// TIA Portal project "uppgift2" (V18) (continued)
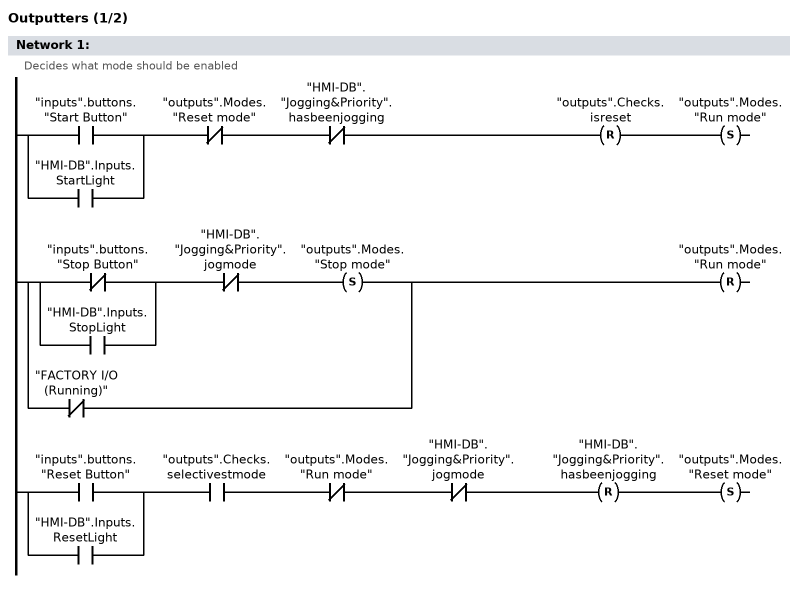
   RUNG wire#powerrail
      Contact( "inputs".buttons."Start Button" )
      wire#w1
      I_Contact( "outputs".Modes."Reset mode" )
      I_Contact( "HMI-DB"."Jogging&Priority".hasbeenjogging )
      R_Coil( "outputs".Checks.isreset )
      S_Coil( "outputs".Modes."Run mode" )
   END_RUNG
   RUNG wire#powerrail
      Contact( "HMI-DB".Inputs.StartLight )
   END_RUNG wire#w1
   RUNG wire#powerrail
      I_Contact( "inputs".buttons."Stop Button" )
      wire#w2
      I_Contact( "HMI-DB"."Jogging&Priority".jogmode )
      S_Coil( "outputs".Modes."Stop mode" )
      wire#w3
      R_Coil( "outputs".Modes."Run mode" )
   END_RUNG
   RUNG wire#powerrail
      Contact( "HMI-DB".Inputs.StopLight )
   END_RUNG wire#w2
   RUNG wire#powerrail
      I_Contact( "FACTORY I/O (Running)" )
   END_RUNG wire#w3
   RUNG wire#powerrail
      Contact( "inputs".buttons."Reset Button" )
      wire#w4
      Contact( "outputs".Checks.selectivestmode )
      I_Contact( "outputs".Modes."Run mode" )
      I_Contact( "HMI-DB"."Jogging&Priority".jogmode )
      R_Coil( "HMI-DB"."Jogging&Priority".hasbeenjogging )
      S_Coil( "outputs".Modes."Reset mode" )
   END_RUNG
   RUNG wire#powerrail
      Contact( "HMI-DB".Inputs.ResetLight )
   END_RUNG wire#w4
   // the same network as SCL:
   IF ("inputs".buttons."Start Button" OR "HMI-DB".Inputs.StartLight) AND NOT "outputs".Modes."Reset mode" AND NOT "HMI-DB"."Jogging&Priority".hasbeenjogging THEN
       "outputs".Checks.isreset := FALSE;
       "outputs".Modes."Run mode" := TRUE;
   END_IF;
   #_w1 := (NOT "inputs".buttons."Stop Button" OR "HMI-DB".Inputs.StopLight) AND NOT "HMI-DB"."Jogging&Priority".jogmode;
   IF #_w1 THEN "outputs".Modes."Stop mode" := TRUE; END_IF;
   IF #_w1 OR NOT "FACTORY I/O (Running)" THEN "outputs".Modes."Run mode" := FALSE; END_IF;
   IF ("inputs".buttons."Reset Button" OR "HMI-DB".Inputs.ResetLight) AND "outputs".Checks.selectivestmode AND NOT "outputs".Modes."Run mode" AND NOT "HMI-DB"."Jogging&Priority".jogmode THEN
       "HMI-DB"."Jogging&Priority".hasbeenjogging := FALSE;
       "outputs".Modes."Reset mode" := TRUE;
   END_IF;
END_REGION

REGION Network 2
   // Turns on the acutators if the correct signal is on
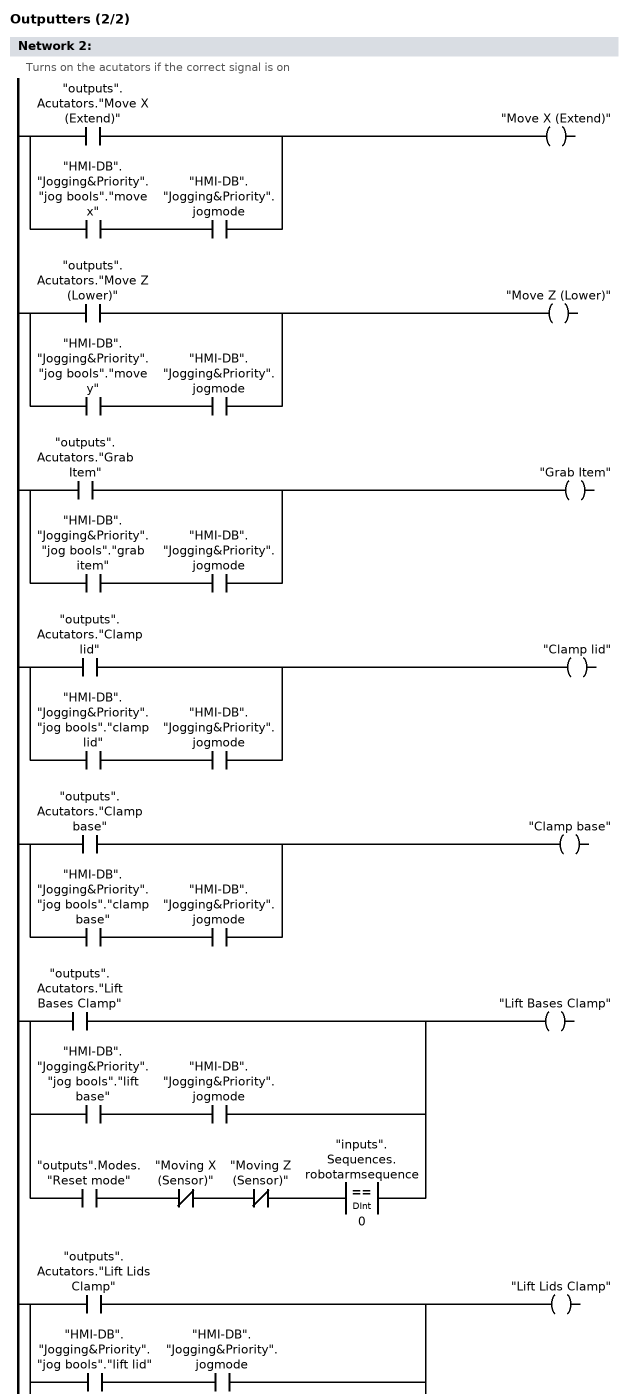
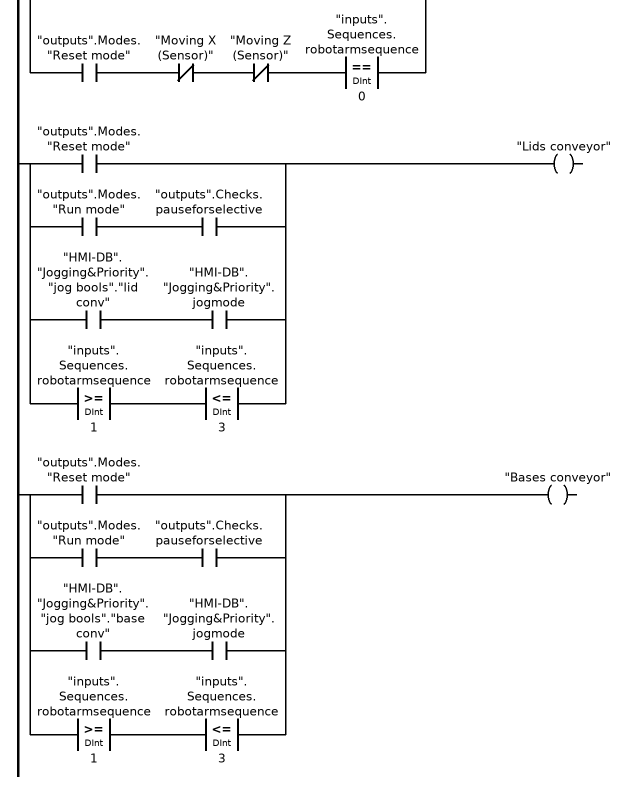
   RUNG wire#powerrail
      Contact( "outputs".Acutators."Move X (Extend)" )
      wire#w1
      Coil( "Move X (Extend)" )
   END_RUNG
   RUNG wire#powerrail
      Contact( "HMI-DB"."Jogging&Priority"."jog bools"."move x" )
      Contact( "HMI-DB"."Jogging&Priority".jogmode )
   END_RUNG wire#w1
   RUNG wire#powerrail
      Contact( "outputs".Acutators."Move Z (Lower)" )
      wire#w2
      Coil( "Move Z (Lower)" )
   END_RUNG
   RUNG wire#powerrail
      Contact( "HMI-DB"."Jogging&Priority"."jog bools"."move y" )
      Contact( "HMI-DB"."Jogging&Priority".jogmode )
   END_RUNG wire#w2
   RUNG wire#powerrail
      Contact( "outputs".Acutators."Grab Item" )
      wire#w3
      Coil( "Grab Item" )
   END_RUNG
   RUNG wire#powerrail
      Contact( "HMI-DB"."Jogging&Priority"."jog bools"."grab item" )
      Contact( "HMI-DB"."Jogging&Priority".jogmode )
   END_RUNG wire#w3
   RUNG wire#powerrail
      Contact( "outputs".Acutators."Clamp lid" )
      wire#w4
      Coil( "Clamp lid" )
   END_RUNG
   RUNG wire#powerrail
      Contact( "HMI-DB"."Jogging&Priority"."jog bools"."clamp lid" )
      Contact( "HMI-DB"."Jogging&Priority".jogmode )
   END_RUNG wire#w4
   RUNG wire#powerrail
      Contact( "outputs".Acutators."Clamp base" )
      wire#w5
      Coil( "Clamp base" )
   END_RUNG
   RUNG wire#powerrail
      Contact( "HMI-DB"."Jogging&Priority"."jog bools"."clamp base" )
      Contact( "HMI-DB"."Jogging&Priority".jogmode )
   END_RUNG wire#w5
   RUNG wire#powerrail
      Contact( "outputs".Acutators."Lift Bases Clamp" )
      wire#w6
      Coil( "Lift Bases Clamp" )
   END_RUNG
   RUNG wire#powerrail
      Contact( "HMI-DB"."Jogging&Priority"."jog bools"."lift base" )
      Contact( "HMI-DB"."Jogging&Priority".jogmode )
   END_RUNG wire#w6
   RUNG wire#powerrail
      Contact( "outputs".Modes."Reset mode" )
      I_Contact( "Moving X (Sensor)" )
      I_Contact( "Moving Z (Sensor)" )
      { S7_Templates := "SrcType := DInt" } EQ_Contact(in1 := "inputs".Sequences.robotarmsequence, in2 := 0)
   END_RUNG wire#w6
   RUNG wire#powerrail
      Contact( "outputs".Acutators."Lift Lids Clamp" )
      wire#w7
      Coil( "Lift Lids Clamp" )
   END_RUNG
   RUNG wire#powerrail
      Contact( "HMI-DB"."Jogging&Priority"."jog bools"."lift lid" )
      Contact( "HMI-DB"."Jogging&Priority".jogmode )
   END_RUNG wire#w7
   RUNG wire#powerrail
      Contact( "outputs".Modes."Reset mode" )
      I_Contact( "Moving X (Sensor)" )
      I_Contact( "Moving Z (Sensor)" )
      { S7_Templates := "SrcType := DInt" } EQ_Contact(in1 := "inputs".Sequences.robotarmsequence, in2 := 0)
   END_RUNG wire#w7
   RUNG wire#powerrail
      Contact( "outputs".Modes."Reset mode" )
      wire#w8
      Coil( "Lids conveyor" )
   END_RUNG
   RUNG wire#powerrail
      Contact( "outputs".Modes."Run mode" )
      Contact( "outputs".Checks.pauseforselective )
   END_RUNG wire#w8
   RUNG wire#powerrail
      Contact( "HMI-DB"."Jogging&Priority"."jog bools"."lid conv" )
      Contact( "HMI-DB"."Jogging&Priority".jogmode )
   END_RUNG wire#w8
   RUNG wire#powerrail
      { S7_Templates := "SrcType := DInt" } GE_Contact(in1 := "inputs".Sequences.robotarmsequence, in2 := 1)
      { S7_Templates := "SrcType := DInt" } LE_Contact(in1 := "inputs".Sequences.robotarmsequence, in2 := 3)
   END_RUNG wire#w8
   RUNG wire#powerrail
      Contact( "outputs".Modes."Reset mode" )
      wire#w9
      Coil( "Bases conveyor" )
   END_RUNG
   RUNG wire#powerrail
      Contact( "outputs".Modes."Run mode" )
      Contact( "outputs".Checks.pauseforselective )
   END_RUNG wire#w9
   RUNG wire#powerrail
      Contact( "HMI-DB"."Jogging&Priority"."jog bools"."base conv" )
      Contact( "HMI-DB"."Jogging&Priority".jogmode )
   END_RUNG wire#w9
   RUNG wire#powerrail
      { S7_Templates := "SrcType := DInt" } GE_Contact(in1 := "inputs".Sequences.robotarmsequence, in2 := 1)
      { S7_Templates := "SrcType := DInt" } LE_Contact(in1 := "inputs".Sequences.robotarmsequence, in2 := 3)
   END_RUNG wire#w9
   // the same network as SCL:
   "Move X (Extend)" := "outputs".Acutators."Move X (Extend)" OR ("HMI-DB"."Jogging&Priority"."jog bools"."move x" AND "HMI-DB"."Jogging&Priority".jogmode);
   "Move Z (Lower)" := "outputs".Acutators."Move Z (Lower)" OR ("HMI-DB"."Jogging&Priority"."jog bools"."move y" AND "HMI-DB"."Jogging&Priority".jogmode);
   "Grab Item" := "outputs".Acutators."Grab Item" OR ("HMI-DB"."Jogging&Priority"."jog bools"."grab item" AND "HMI-DB"."Jogging&Priority".jogmode);
   "Clamp lid" := "outputs".Acutators."Clamp lid" OR ("HMI-DB"."Jogging&Priority"."jog bools"."clamp lid" AND "HMI-DB"."Jogging&Priority".jogmode);
   "Clamp base" := "outputs".Acutators."Clamp base" OR ("HMI-DB"."Jogging&Priority"."jog bools"."clamp base" AND "HMI-DB"."Jogging&Priority".jogmode);
   "Lift Bases Clamp" := "outputs".Acutators."Lift Bases Clamp" OR ("HMI-DB"."Jogging&Priority"."jog bools"."lift base" AND "HMI-DB"."Jogging&Priority".jogmode) OR ("outputs".Modes."Reset mode" AND NOT "Moving X (Sensor)" AND NOT "Moving Z (Sensor)" AND ("inputs".Sequences.robotarmsequence = 0));
   "Lift Lids Clamp" := "outputs".Acutators."Lift Lids Clamp" OR ("HMI-DB"."Jogging&Priority"."jog bools"."lift lid" AND "HMI-DB"."Jogging&Priority".jogmode) OR ("outputs".Modes."Reset mode" AND NOT "Moving X (Sensor)" AND NOT "Moving Z (Sensor)" AND ("inputs".Sequences.robotarmsequence = 0));
   "Lids conveyor" := "outputs".Modes."Reset mode" OR ("outputs".Modes."Run mode" AND "outputs".Checks.pauseforselective) OR ("HMI-DB"."Jogging&Priority"."jog bools"."lid conv" AND "HMI-DB"."Jogging&Priority".jogmode) OR (("inputs".Sequences.robotarmsequence >= 1) AND ("inputs".Sequences.robotarmsequence <= 3));
   "Bases conveyor" := "outputs".Modes."Reset mode" OR ("outputs".Modes."Run mode" AND "outputs".Checks.pauseforselective) OR ("HMI-DB"."Jogging&Priority"."jog bools"."base conv" AND "HMI-DB"."Jogging&Priority".jogmode) OR (("inputs".Sequences.robotarmsequence >= 1) AND ("inputs".Sequences.robotarmsequence <= 3));
END_REGION
END_FUNCTION

// folder: lids/bases

FUNCTION "lids" : Void   // FC3, LAD
{ S7_Optimized_Access := 'TRUE' }
VERSION : 0.1
// Controls the lid clamp and lift and controls when the robots sequence should start
   VAR_TEMP   // added for the SCL form of the ladder/FBD networks
      _w1 : Bool;
   END_VAR
BEGIN

REGION Network 1
   // Runs the emitter if sequence is 0 and lids vision doesnt detect any lid
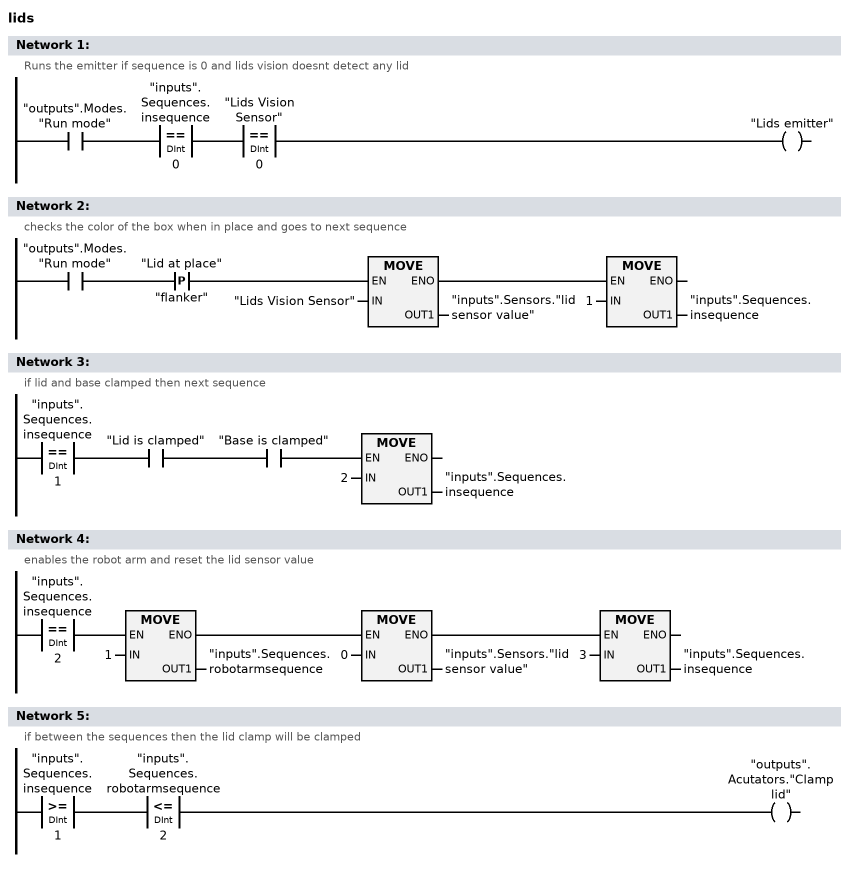
   RUNG wire#powerrail
      Contact( "outputs".Modes."Run mode" )
      { S7_Templates := "SrcType := DInt" } EQ_Contact(in1 := "inputs".Sequences.insequence, in2 := 0)
      { S7_Templates := "SrcType := DInt" } EQ_Contact(in1 := "Lids Vision Sensor", in2 := 0)
      Coil( "Lids emitter" )
   END_RUNG
   // the same network as SCL:
   "Lids emitter" := "outputs".Modes."Run mode" AND ("inputs".Sequences.insequence = 0) AND ("Lids Vision Sensor" = 0);
END_REGION

REGION Network 2
   // checks the color of the box when in place and goes to next sequence
   RUNG wire#powerrail
      Contact( "outputs".Modes."Run mode" )
      P_Contact(operand := "Lid at place", bit := "flanker")
      Move(in := "Lids Vision Sensor", out1 => "inputs".Sensors."lid sensor value")
      Move(in := 1, out1 => "inputs".Sequences.insequence)
   END_RUNG
   // the same network as SCL:
   #_w1 := "outputs".Modes."Run mode" AND "Lid at place" AND NOT "flanker";   // rising edge of "Lid at place"
   "flanker" := "Lid at place";
   IF #_w1 THEN
       "inputs".Sensors."lid sensor value" := "Lids Vision Sensor";
       "inputs".Sequences.insequence := 1;
   END_IF;
END_REGION

REGION Network 3
   // if lid and base clamped then next sequence
   RUNG wire#powerrail
      { S7_Templates := "SrcType := DInt" } EQ_Contact(in1 := "inputs".Sequences.insequence, in2 := 1)
      Contact( "Lid is clamped" )
      Contact( "Base is clamped" )
      Move(in := 2, out1 => "inputs".Sequences.insequence)
   END_RUNG
   // the same network as SCL:
   IF ("inputs".Sequences.insequence = 1) AND "Lid is clamped" AND "Base is clamped" THEN
       "inputs".Sequences.insequence := 2;
   END_IF;
END_REGION

REGION Network 4
   // enables the robot arm and reset the lid sensor value
   RUNG wire#powerrail
      { S7_Templates := "SrcType := DInt" } EQ_Contact(in1 := "inputs".Sequences.insequence, in2 := 2)
      Move(in := 1, out1 => "inputs".Sequences.robotarmsequence)
      Move(in := 0, out1 => "inputs".Sensors."lid sensor value")
      Move(in := 3, out1 => "inputs".Sequences.insequence)
   END_RUNG
   // the same network as SCL:
   IF "inputs".Sequences.insequence = 2 THEN
       "inputs".Sequences.robotarmsequence := 1;
       "inputs".Sensors."lid sensor value" := 0;
       "inputs".Sequences.insequence := 3;
   END_IF;
END_REGION

REGION Network 5
   // if between the sequences then the lid clamp will be clamped
   RUNG wire#powerrail
      { S7_Templates := "SrcType := DInt" } GE_Contact(in1 := "inputs".Sequences.insequence, in2 := 1)
      { S7_Templates := "SrcType := DInt" } LE_Contact(in1 := "inputs".Sequences.robotarmsequence, in2 := 2)
      Coil( "outputs".Acutators."Clamp lid" )
   END_RUNG
   // the same network as SCL:
   "outputs".Acutators."Clamp lid" := ("inputs".Sequences.insequence >= 1) AND ("inputs".Sequences.robotarmsequence <= 2);
END_REGION
END_FUNCTION

FUNCTION "base" : Void   // FC6, LAD
{ S7_Optimized_Access := 'TRUE' }
VERSION : 0.1
// Controls the base clamp and lift
   VAR_TEMP   // added for the SCL form of the ladder/FBD networks
      _w1 : Bool;
   END_VAR
BEGIN

REGION Network 1
   // If base sequence is 0 and no item is at base at place sensor, then the emitter will run
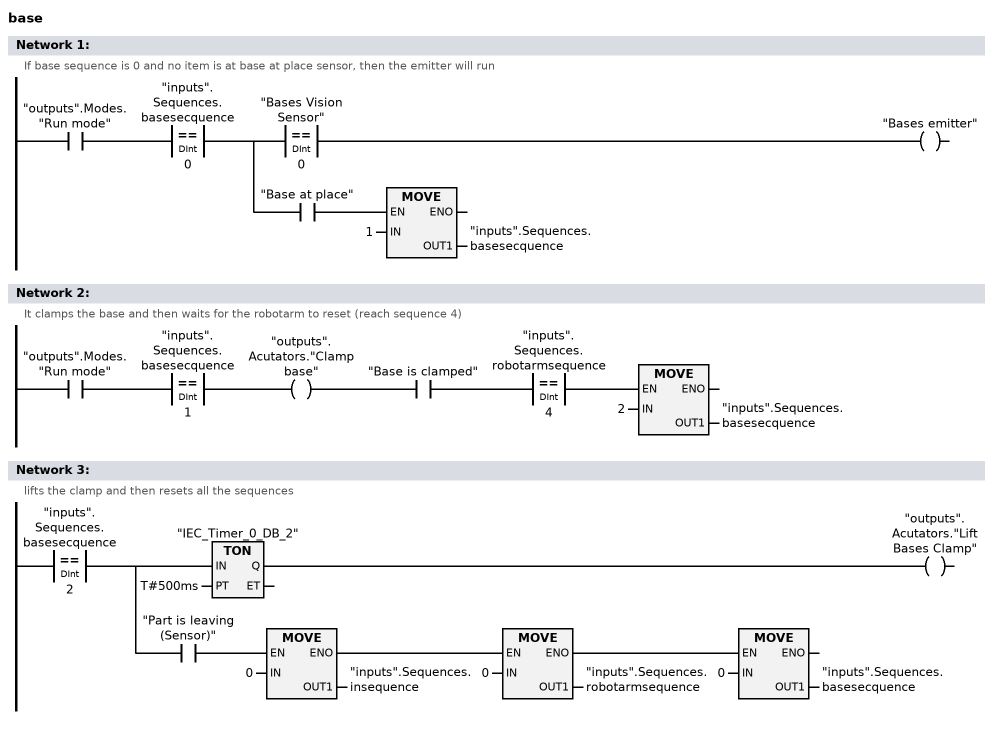
   RUNG wire#powerrail
      Contact( "outputs".Modes."Run mode" )
      { S7_Templates := "SrcType := DInt" } EQ_Contact(in1 := "inputs".Sequences.basesecquence, in2 := 0)
      wire#w1
      { S7_Templates := "SrcType := DInt" } EQ_Contact(in1 := "Bases Vision Sensor", in2 := 0)
      Coil( "Bases emitter" )
   END_RUNG
   RUNG wire#w1
      Contact( "Base at place" )
      Move(in := 1, out1 => "inputs".Sequences.basesecquence)
   END_RUNG
   // the same network as SCL:
   #_w1 := "outputs".Modes."Run mode" AND ("inputs".Sequences.basesecquence = 0);
   "Bases emitter" := #_w1 AND ("Bases Vision Sensor" = 0);
   IF #_w1 AND "Base at place" THEN "inputs".Sequences.basesecquence := 1; END_IF;
END_REGION

REGION Network 2
   // It clamps the base and then waits for the robotarm to reset (reach sequence 4)
   RUNG wire#powerrail
      Contact( "outputs".Modes."Run mode" )
      { S7_Templates := "SrcType := DInt" } EQ_Contact(in1 := "inputs".Sequences.basesecquence, in2 := 1)
      Coil( "outputs".Acutators."Clamp base" )
      Contact( "Base is clamped" )
      { S7_Templates := "SrcType := DInt" } EQ_Contact(in1 := "inputs".Sequences.robotarmsequence, in2 := 4)
      Move(in := 2, out1 => "inputs".Sequences.basesecquence)
   END_RUNG
   // the same network as SCL:
   "outputs".Acutators."Clamp base" := "outputs".Modes."Run mode" AND ("inputs".Sequences.basesecquence = 1);
   IF "outputs".Acutators."Clamp base" AND "Base is clamped" AND ("inputs".Sequences.robotarmsequence = 4) THEN
       "inputs".Sequences.basesecquence := 2;
   END_IF;
END_REGION

REGION Network 3
   // lifts the clamp and then resets all the sequences
   #_w1 := "inputs".Sequences.basesecquence = 2;
   "IEC_Timer_0_DB_2".TON(IN := #_w1, PT := T#500ms);
   "outputs".Acutators."Lift Bases Clamp" := "IEC_Timer_0_DB_2".Q;
   IF #_w1 AND "Part is leaving (Sensor)" THEN
       "inputs".Sequences.insequence := 0;
       "inputs".Sequences.robotarmsequence := 0;
       "inputs".Sequences.basesecquence := 0;
   END_IF;
END_REGION
END_FUNCTION

(* ===== HMI "HMI_RT_1" =====
system functions are stored by id; their names below are inferred from use
connection "PLC": ETHERNET, S7_1200_OMS
connection "HMI_Connection_1": ETHERNET, S7_1500_OMS

HMI tags "Default tag table"
   "Input1" : Bool = PLC "Start Light" AT %Q1.0, 1 s
   "Input2" : Bool = PLC hmistop AT %I2.2, 1 s
   "Input3" : Bool = PLC hmireset AT %I2.3, 1 s
   "inputs_buttons_Start Button" : Bool = PLC inputs.buttons."Start Button", 1 s
   "HMI-DB_Inputs_StartLight" : Bool = PLC "HMI-DB".Inputs.StartLight, 1 s
   "HMI-DB_Inputs_StopLight" : Bool = PLC "HMI-DB".Inputs.StopLight, 1 s
   "HMI-DB_Inputs_ResetLight" : Bool = PLC "HMI-DB".Inputs.ResetLight, 1 s
   "HMI-DB_Internal_jogmode" : Bool = PLC "HMI-DB".Jogging&Priority.jogmode, 1 s
   "HMI-DB_Internal_jogthings_move x" : Bool = PLC "HMI-DB".Jogging&Priority."jog bools"."move x", 1 s
   "HMI-DB_Internal_jogthings_move y" : Bool = PLC "HMI-DB".Jogging&Priority."jog bools"."move y", 1 s
   "HMI-DB_Internal_jogthings_grab item" : Bool = PLC "HMI-DB".Jogging&Priority."jog bools"."grab item", 1 s
   "HMI-DB_Internal_jogthings_clamp lid" : Bool = PLC "HMI-DB".Jogging&Priority."jog bools"."clamp lid", 1 s
   "HMI-DB_Internal_jogthings_clamp base" : Bool = PLC "HMI-DB".Jogging&Priority."jog bools"."clamp base", 1 s
   "HMI-DB_Internal_jogthings_lift base" : Bool = PLC "HMI-DB".Jogging&Priority."jog bools"."lift base", 1 s
   "HMI-DB_Internal_jogthings_lift lid" : Bool = PLC "HMI-DB".Jogging&Priority."jog bools"."lift lid", 1 s
   "HMI-DB_Internal_jogthings_lid conv" : Bool = PLC "HMI-DB".Jogging&Priority."jog bools"."lid conv", 1 s
   "HMI-DB_Internal_jogthings_base conv" : Bool = PLC "HMI-DB".Jogging&Priority."jog bools"."base conv", 1 s
   "HMI-DB_Internal_jogthings_lampor" : Bool = PLC "HMI-DB".Jogging&Priority."jog bools".lampor, 1 s
   "movexlight" : Bool = PLC "Moving X (Sensor)" AT %I1.4, 1 s
   "moveylight" : Bool = PLC "Moving Z (Sensor)" AT %I1.5, 1 s
   "lidclampedlight" : Bool = PLC "Lid is clamped" AT %I1.0, 1 s
   "baseisclamplight" : Bool = PLC "Base is clamped" AT %I0.7, 1 s
   "itemdetectlight" : Bool = PLC "Item detected" AT %I1.1, 1 s
   "lidatplacelight" : Bool = PLC "Lid at place" AT %I0.6, 1 s
   "baseatplacelight" : Bool = PLC "Base at place" AT %I0.5, 1 s
   "partisleavinglight" : Bool = PLC "Part is leaving (Sensor)" AT %I1.2, 1 s
   "lidisleavinglight" : Bool = PLC IEC_Counter_0_DB_2.CD AT %I1.6, 1 s
   "outputs_Run mode" : Bool = PLC outputs.Modes."Run mode", 1 s
   "outputs_Stop mode" : Bool = PLC outputs.Modes."Stop mode", 1 s
   "outputs_Reset mode" : Bool = PLC outputs.Modes."Reset mode", 1 s
   "outputs_blue lids" : Int = PLC outputs.BoxesCounters."blue lids", 1 s
   "Lift Lids Clamp" : Bool = PLC "Lift Lids Clamp" AT %Q0.7, 1 s
   "baselift clamp limit" : Bool = PLC "baselift clamp limit" AT %I1.7, 1 s
   "lift lids clamp limit" : Bool = PLC "lids lift clamp limit" AT %I1.6, 1 s
   "outputs_green lids" : Int = PLC outputs.BoxesCounters."green lids", 1 s
   "RESET!!!!!!!!!" : Bool = PLC "HMI-DB".Jogging&Priority.resetdelivered, 1 s
   "outputs_blue bases" : Int = PLC outputs.BoxesCounters."blue bases", 1 s
   "outputs_green bases" : Int = PLC outputs.BoxesCounters."green bases", 1 s
   "outputs_blue boxs" : Int = PLC outputs.BoxesCounters."blue boxs", 1 s
   "outputs_green boxs" : Int = PLC outputs.BoxesCounters."green boxs", 1 s
   "outputs_greenblue box" : Int = PLC outputs.BoxesCounters."greenblue box", 1 s
   "outputs_bluegreen box" : Int = PLC outputs.BoxesCounters."bluegreen box", 1 s
   "outputs_selectivestmode" : Bool = PLC outputs.Checks.selectivestmode, 1 s
   "HMI-DB_Internal_hmipriority" : Bool = PLC "HMI-DB".Jogging&Priority.hmipriority, 1 s
   "HMI-DB_Internal_hmiprioritystate" : Bool = PLC "HMI-DB".Jogging&Priority.hmiprioritystate, 1 s
   "outputs_toproduceeeee" : Int = PLC outputs.Hmi-Producer.toproduce, 1 s
   "outputs_producedboxes" : Int = PLC outputs.Hmi-Producer.producedboxes, 1 s
   "outputs_robotarmsequence" : DInt = PLC inputs.Sequences.robotarmsequence, 1 s
   "inputs_basesecquence" : DInt = PLC inputs.Sequences.basesecquence, 1 s
   "inputs_insequence" : DInt = PLC inputs.Sequences.insequence, 1 s
   "Counter" : DInt = PLC Counter AT %QD30, 1 s
   "outputs_totalpartscounter" : Int = PLC outputs.BoxesCounters.totalpartscounter, 1 s
   "outputs_Move X (Extend)" : Bool = PLC outputs.Acutators."Move X (Extend)", 1 s
   "outputs_Move Z (Lower)" : Bool = PLC outputs.Acutators."Move Z (Lower)", 1 s
   "outputs_Grab Item" : Bool = PLC outputs.Acutators."Grab Item", 1 s
   "outputs_Clamp base" : Bool = PLC outputs.Acutators."Clamp base", 1 s
   "outputs_Clamp lid" : Bool = PLC outputs.Acutators."Clamp lid", 1 s
   "outputs_Lift Bases Clamp" : Bool = PLC outputs.Acutators."Lift Bases Clamp", 1 s
   "outputs_Lift Lids Clamp" : Bool = PLC outputs.Acutators."Lift Lids Clamp", 1 s
   "Lids conveyor" : Bool = PLC "Lids conveyor" AT %Q1.3, 1 s
   "Bases conveyor" : Bool = PLC "Bases conveyor" AT %Q1.4, 1 s
   "inputs_green light" : Bool = PLC inputs."green light", 1 s
   "outputs_RESETBUTTONHMI" : Bool = PLC outputs.RESETBUTTONHMI, 1 s
   "Move X (Extend)" : Bool = PLC "Move X (Extend)" AT %Q0.0, 1 s
   "Move Z (Lower)" : Bool = PLC "Move Z (Lower)" AT %Q0.1, 1 s
   "Grab Item" : Bool = PLC "Grab Item" AT %Q0.2, 1 s
   "Clamp lid" : Bool = PLC "Clamp lid" AT %Q0.4, 1 s
   "Clamp base" : Bool = PLC "Clamp base" AT %Q0.3, 1 s
   "Lift Bases Clamp" : Bool = PLC "Lift Bases Clamp" AT %Q0.6, 1 s

Template "Template_1" 800x480
   TextField "Template_Text field_1" at 328,22 size 152x43; Text 'amorbus'
   SymbolicIOField "Template_Symbolic I/O field_1" at 108,22 size 170x32; TextOff '0'; TextOn '1'
   Button "Template_Button_1" at 126,248 size 96x32; TextOff 'staaaart'
   Button "Template_Button_2" at 302,248 size 96x32; TextOff 'stop'
   Button "Template_Button_3" at 474,248 size 96x32; TextOff 'reset'
   Button "Template_Button_4" at 302,404 size 96x32; TextOff 'jog it'

screen "root screen" 800x480
   TextField "Template_Text field_1" at 328,22 size 191x43; Text 'Main menu'
   Button "Template_Button_1" at 626,84 size 161x78; TextOff 'Start'
      on Press: SetBit("HMI-DB_Inputs_StartLight")
      on Release: ResetBit("HMI-DB_Inputs_StartLight")
      Appearance <- "outputs_Run mode"
   Button "Template_Button_2" at 626,173 size 161x78; TextOff 'Stop'
      on Press: SetBit("HMI-DB_Inputs_StopLight")
      on Release: ResetBit("HMI-DB_Inputs_StopLight")
      Appearance <- "outputs_Stop mode"
   Button "Template_Button_3" at 626,263 size 161x78; TextOff 'Reset'
      on Press: SetBit("HMI-DB_Inputs_ResetLight")
      on Release: ResetBit("HMI-DB_Inputs_ResetLight")
      Appearance <- "outputs_Reset mode"
   Button "Button_1" at 625,389 size 160x32; TextOff 'Next page'
      on Click: ActivateScreen("joggyes", 0)
   Button "Button_2" at 344,309 size 96x32; TextOff 'Auto'
      Appearance <- "HMI-DB_Internal_hmipriority"
      Visibility <- "HMI-DB_Internal_hmipriority"
      on Click: InvertBit("HMI-DB_Internal_hmipriority")
   Button "Button_3" at 344,309 size 96x32; TextOff 'Selective'
      Visibility <- "HMI-DB_Internal_hmipriority"
      Appearance <- "HMI-DB_Internal_hmipriority"
      on Click: InvertBit("HMI-DB_Internal_hmipriority")
   Button "Button_4" at 323,388 size 139x32; TextOff 'HMI Priority'
      Appearance <- "HMI-DB_Internal_hmiprioritystate"
      on Click: InvertBit("HMI-DB_Internal_hmiprioritystate")
   Bar "Bar_1" at 32,220 size 80x171; MinimumValue 0; MaximumValue 4
      ProcessValue <- "outputs_robotarmsequence"
   Bar "Bar_2" at 128,220 size 80x171; MinimumValue 0; MaximumValue 3
      ProcessValue <- "inputs_insequence"
   Bar "Bar_3" at 223,220 size 80x171; MinimumValue 0; MaximumValue 3
      ProcessValue <- "inputs_basesecquence"
   TextField "Text field_1" at 43,424 size 42x23; Text 'Arm'
   TextField "Text field_2" at 143,424 size 32x23; Text 'Lid'
   TextField "Text field_3" at 237,424 size 48x23; Text 'Base'
   TextField "Text field_4" at 28,173 size 211x23; Text 'Process status percent'

screen "joggyes" 800x480
   Button "Button_1" at 29,402 size 209x32; TextOff 'previous screen'
      on Click: ActivateScreen("root screen", 0)
   Button "Button_2" at 20,45 size 117x32; TextOff 'move x'
      on Press: SetBit("HMI-DB_Internal_jogthings_move x")
      on Release: ResetBit("HMI-DB_Internal_jogthings_move x")
      Appearance <- "Move X (Extend)"
   Button "Button_3" at 22,109 size 114x32; TextOff 'move y'
      on Press: SetBit("HMI-DB_Internal_jogthings_move y")
      on Release: ResetBit("HMI-DB_Internal_jogthings_move y")
      Appearance <- "Move Z (Lower)"
   Button "Button_4" at 22,173 size 114x32; TextOff 'grab item'
      on Press: SetBit("HMI-DB_Internal_jogthings_grab item")
      on Release: ResetBit("HMI-DB_Internal_jogthings_grab item")
      Appearance <- "Grab Item"
   Button "Button_5" at 21,239 size 116x32; TextOff 'clamp lid'
      on Press: SetBit("HMI-DB_Internal_jogthings_clamp lid")
      on Release: ResetBit("HMI-DB_Internal_jogthings_clamp lid")
      Appearance <- "Clamp lid"
   Button "Button_6" at 19,295 size 120x32; TextOff 'clamp base'
      on Press: SetBit("HMI-DB_Internal_jogthings_clamp base")
      on Release: ResetBit("HMI-DB_Internal_jogthings_clamp base")
      Appearance <- "Clamp base"
   Button "Button_7" at 252,48 size 110x32; TextOff 'lift base'
      on Press: SetBit("HMI-DB_Internal_jogthings_lift base")
      on Release: ResetBit("HMI-DB_Internal_jogthings_lift base")
      Appearance <- "Lift Bases Clamp"
   Button "Button_8" at 251,112 size 113x32; TextOff 'lift lid'
      on Press: SetBit("HMI-DB_Internal_jogthings_lift lid")
      on Release: ResetBit("HMI-DB_Internal_jogthings_lift lid")
      Appearance <- "Lift Lids Clamp"
   Button "Button_9" at 251,176 size 112x32; TextOff 'lid conv'
      on Press: SetBit("HMI-DB_Internal_jogthings_lid conv")
      on Release: ResetBit("HMI-DB_Internal_jogthings_lid conv")
      Appearance <- "Lids conveyor"
   Button "Button_10" at 250,242 size 114x32; TextOff 'base conv'
      on Press: SetBit("HMI-DB_Internal_jogthings_base conv")
      on Release: ResetBit("HMI-DB_Internal_jogthings_base conv")
      Appearance <- "Bases conveyor"
   Circle "Circle_1" at 680,5 size 25x25
      Appearance <- "movexlight"
   TextField "Text field_1" at 497,3 size 87x23; Text 'Moving X'
   TextField "Text field_2" at 497,39 size 87x23; Text 'Moving Y'
   TextField "Text field_3" at 485,76 size 112x23; Text 'Lid is clamp'
   TextField "Text field_4" at 477,111 size 128x23; Text 'Base is clamp'
   TextField "Text field_5" at 485,145 size 112x23; Text 'Item detect'
   TextField "Text field_6" at 485,178 size 111x23; Text 'Lid at place'
   TextField "Text field_7" at 478,209 size 126x23; Text 'base at place'
   TextField "Text field_8" at 478,240 size 125x23; Text 'part is leavin'
   TextField "Text field_9" at 486,275 size 110x23; Text 'lid is leavin'
   Button "Button_11" at 251,296 size 113x32; TextOff 'test lampor'
      on Press: SetBit("HMI-DB_Internal_jogthings_lampor")
      on Release: ResetBit("HMI-DB_Internal_jogthings_lampor")
      Appearance <- "Input1"
   Circle "Circle_2" at 680,41 size 25x25
      Appearance <- "moveylight"
   Circle "Circle_3" at 680,76 size 25x25
      Appearance <- "lidclampedlight"
   Circle "Circle_4" at 680,113 size 25x25
      Appearance <- "baseisclamplight"
   Circle "Circle_5" at 680,145 size 25x25
      Appearance <- "itemdetectlight"
   Circle "Circle_6" at 680,180 size 25x25
      Appearance <- "lidatplacelight"
   Circle "Circle_7" at 680,212 size 25x25
      Appearance <- "baseatplacelight"
   Circle "Circle_8" at 680,245 size 25x25
      Appearance <- "partisleavinglight"
   Circle "Circle_9" at 680,278 size 25x25
      Appearance <- "lidisleavinglight"
   Button "Button_12" at 373,401 size 124x32; TextOff 'jogmode'
      on Click: InvertBit("HMI-DB_Internal_jogmode")
      Appearance <- "HMI-DB_Internal_jogmode"
   Button "Button_13" at 680,401 size 96x32; TextOff 'Next'
      on Click: ActivateScreen("orderscreen", 0)
   TextField "Text field_10" at 476,309 size 129x23; Text 'lift lids clamp'
   TextField "Text field_11" at 471,344 size 139x23; Text 'lift base clamp'
   Circle "Circle_10" at 680,311 size 25x25
      Appearance <- "lift lids clamp limit"
   Circle "Circle_11" at 680,344 size 25x25
      Appearance <- "baselift clamp limit"

screen "orderscreen" 800x480
   TextField "Text field_1" at 7,324 size 69x18; Text 'Blue lids:'
   TextField "Text field_3" at 0,379 size 79x18; Text 'Green lids:'
   TextField "Text field_5" at 202,324 size 77x18; Text 'Blue base:'
   TextField "Text field_7" at 195,379 size 87x18; Text 'Green base:'
   TextField "Text field_9" at 396,324 size 71x18; Text 'Blue box:'
   TextField "Text field_11" at 389,379 size 81x18; Text 'Green box:'
   TextField "Text field_13" at 575,324 size 117x18; Text 'Green-blue box:'
   TextField "Text field_15" at 576,379 size 117x18; Text 'Blue-green box:'
   IOField "I/O field_1" at 104,320 size 76x32; FormatPattern 9999
      ProcessValue <- "outputs_blue lids"
   IOField "I/O field_2" at 105,375 size 75x32; FormatPattern 9999
      ProcessValue <- "outputs_green lids"
   IOField "I/O field_3" at 299,320 size 75x32; FormatPattern 9999
      ProcessValue <- "outputs_blue bases"
   IOField "I/O field_4" at 299,375 size 76x32; FormatPattern 9999
      ProcessValue <- "outputs_green bases"
   IOField "I/O field_5" at 482,320 size 76x32; FormatPattern 9999
      ProcessValue <- "outputs_blue boxs"
   IOField "I/O field_6" at 482,375 size 77x32; FormatPattern 9999
      ProcessValue <- "outputs_green boxs"
   IOField "I/O field_7" at 710,320 size 75x32; FormatPattern 9999
      ProcessValue <- "outputs_greenblue box"
   IOField "I/O field_8" at 710,375 size 75x32; FormatPattern 9999
      ProcessValue <- "outputs_bluegreen box"
   Button "Button_1" at 46,417 size 209x32; TextOff 'Previous screen'
      on Click: ActivateScreen("joggyes", 0)
   TextField "Text field_2" at 263,0 size 231x47; Text 'Box orderer'
   IOField "I/O field_9" at 199,106 size 145x77; FormatPattern 9999
      ProcessValue <- "outputs_toproduceeeee"
   Button "Button_2" at 295,216 size 145x32; TextOff 'reset counters'
      on Press: SetBit("outputs_RESETBUTTONHMI")
      on Release: ResetBit("outputs_RESETBUTTONHMI")
   TextField "Text field_4" at 199,74 size 130x23; Text 'Order amount'
   IOField "I/O field_10" at 389,106 size 145x77; FormatPattern 9999
      ProcessValue <- "outputs_producedboxes"
   TextField "Text field_6" at 389,74 size 177x23; Text 'has been delivered'
   TextField "Text field_8" at 592,263 size 92x18; Text 'Total boxes:'
   IOField "I/O field_11" at 710,261 size 76x32; FormatPattern 9999
      ProcessValue <- "outputs_totalpartscounter"
*)